// Mitsubishi GX Works2 project: 40国轩高温2次注液尝试优化   PLC: Q06UDEH (continued)

Lifter40204(ShuttleCarInOut:=LifterIO40204);	(*2线升降台*)
LifterIO40204.xCylinder:=1;
Y240:=LifterIO40204.xCW;					
Y241:=LifterIO40204.xCCW;					
LifterIO40204.xForward:=M549;					
LifterIO40204.xBackward:=M550;					
ShuttleCarCurrentPosition(X45 OR X44,X44,X45,FALSE,LifterIO40204.iCurrentPos);					
M647:=LifterIO40204.xOvertimeAlarm ;					
LifterIO40204.diDeviceID:=40204;					

Lifter40205(ShuttleCarInOut:=LifterIO40205);		(*3线升降台*)
LifterIO40205.xCylinder:=1;			
Y242:=LifterIO40205.xCW;					
Y243:=LifterIO40205.xCCW;					
LifterIO40205.xForward:=M551;					
LifterIO40205.xBackward:=M552;					
ShuttleCarCurrentPosition(X47 OR X46,X47,X46,FALSE,LifterIO40205.iCurrentPos);					
M648:=LifterIO40205.xOvertimeAlarm ;					
LifterIO40205.diDeviceID:=40205;					

Lifter40206(ShuttleCarInOut:=LifterIO40206);	(*4线升降台*)	
LifterIO40206.xCylinder:=1;			
Y276:=LifterIO40206.xCW;					
Y244:=LifterIO40206.xCCW;					
LifterIO40206.xForward:=M553;					
LifterIO40206.xBackward:=M554;					
ShuttleCarCurrentPosition(X49 OR X48,X48,X49,FALSE,LifterIO40206.iCurrentPos);					
M649:=LifterIO40206.xOvertimeAlarm ;					
LifterIO40206.diDeviceID:=40206;					

Lifter40207(ShuttleCarInOut:=LifterIO40207);	(*高温入库顶起机构*)	
LifterIO40207.xCylinder:=1;			
Y256:=LifterIO40207.xCW;					
Y257:=LifterIO40207.xCCW;					
LifterIO40207.xForward:=M556;					
LifterIO40207.xBackward:=M583;					
ShuttleCarCurrentPosition(X66 OR X65,X66,X65,FALSE,LifterIO40207.iCurrentPos);					
LifterIO40206.diDeviceID:=40207;
M651:=LifterIO40207.xOvertimeAlarm ;	

Lifter40208(ShuttleCarInOut:=LifterIO40208);	(*高温出库顶起机构*)	
LifterIO40208.xCylinder:=1;			
Y25A:=LifterIO40208.xCW;					
Y25B:=LifterIO40208.xCCW;					
LifterIO40208.xForward:=M558;					
LifterIO40208.xBackward:=M584;					
ShuttleCarCurrentPosition(X6A OR X69,X6A,X69,FALSE,LifterIO40208.iCurrentPos);					
LifterIO40206.diDeviceID:=40208;	
M653:=LifterIO40206.xOvertimeAlarm ;		

Switch40301(ConveyorEntryIO:=ConveyorIO40101 ,ConveyorExitIO:=ConveyorIO40102 ,SwitchIO:=SwitchIO40301);(*高温入库*)
SwitchIO40301.xLiftCylinderRetractDetect:=X64;							
SwitchIO40301.xLiftCylinderExtendDetect:=X63;							
Y254:=SwitchIO40301.xLiftCylinderExtend;							
SwitchIO40301.xLiftCylinderExtendButton:=M555;	
SwitchIO40301.xLiftCylinderRetractButton:=NOT M555;						
M650:=SwitchIO40301.xOvertimeAlarm ;							

(*Switch40302(ConveyorEntryIO:=ConveyorIO40103 ,ConveyorExitIO:=ConveyorIO40104 ,SwitchIO:=SwitchIO40302);*)(*高温入库里面*)(*
SwitchIO40302.xLiftCylinderRetractDetect:=X66;						
SwitchIO40302.xLiftCylinderExtendDetect:=X65;		*)										
						

Switch40303(ConveyorEntryIO:=ConveyorIO40106 ,ConveyorExitIO:=ConveyorIO40109 ,SwitchIO:=SwitchIO40303);(*高温出库*)
SwitchIO40303.xLiftCylinderExtendInit:=1;
SwitchIO40303.xLiftCylinderRetractDetect:=X68;							
SwitchIO40303.xLiftCylinderExtendDetect:=X67;							
Y258:=SwitchIO40303.xLiftCylinderExtend;							
SwitchIO40303.xLiftCylinderExtendButton:=M557;	
SwitchIO40303.xLiftCylinderRetractButton:=NOT M557;						
M652:=SwitchIO40303.xOvertimeAlarm ;							
SwitchIO40303.xLiftCylinderExtendInit:=1;

Switch40304(ConveyorEntryIO:=ConveyorIO40108 ,ConveyorExitIO:=ConveyorIO40107 ,SwitchIO:=SwitchIO40304);(*高温出库里面*)
SwitchIO40304.xLiftCylinderExtendInit:=1;
SwitchIO40304.xLiftCylinderRetractDetect:=X6A;	(*顶起部分单独写了*)						
SwitchIO40304.xLiftCylinderExtendDetect:=X69;											
SwitchIO40304.xLiftCylinderExtendInit:=1;						

Switch40305(ConveyorEntryIO:=ConveyorIO40114 ,ConveyorExitIO:=ConveyorIO40110 ,SwitchIO:=SwitchIO40305);(*1线上层*)
SwitchIO40305.xLiftCylinderRetractDetect:=X6C;							
SwitchIO40305.xLiftCylinderExtendDetect:=X6B;							
Y25C:=SwitchIO40305.xLiftCylinderExtend;							
Y270:=SwitchIO40305.xExitBarCylinderRetract;							
SwitchIO40305.xLiftCylinderExtendButton:=M559;	
SwitchIO40305.xLiftCylinderRetractButton:=NOT M559;						
SwitchIO40305.xExitBarCylinderRetractButton:=M560;							
M654:=SwitchIO40305.xOvertimeAlarm ;							

Switch40306(ConveyorEntryIO:=ConveyorIO40112 ,ConveyorExitIO:=ConveyorIO40113 ,SwitchIO:=SwitchIO40306);(*2线上层*)
SwitchIO40306.xLiftCylinderRetractDetect:=X6E;							
SwitchIO40306.xLiftCylinderExtendDetect:=X6D;							
Y25E:=SwitchIO40306.xLiftCylinderExtend;							
Y279:=SwitchIO40306.xExitBarCylinderRetract;							
SwitchIO40306.xLiftCylinderExtendButton:=M561;	
SwitchIO40306.xLiftCylinderRetractButton:=NOT M561;						
SwitchIO40306.xExitBarCylinderRetractButton:=M562;							
M655:=SwitchIO40306.xOvertimeAlarm ;							

Switch40307(ConveyorEntryIO:=ConveyorIO40115 ,ConveyorExitIO:=ConveyorIO40116 ,SwitchIO:=SwitchIO40307);(*3线上层*)
SwitchIO40307.xLiftCylinderRetractDetect:=X70;							
SwitchIO40307.xLiftCylinderExtendDetect:=X6F;							
Y260:=SwitchIO40307.xLiftCylinderExtend;							
Y27A:=SwitchIO40307.xExitBarCylinderRetract;							
SwitchIO40307.xLiftCylinderExtendButton:=M563;	
SwitchIO40307.xLiftCylinderRetractButton:=NOT M563;						
SwitchIO40307.xExitBarCylinderRetractButton:=M564;							
M656:=SwitchIO40307.xOvertimeAlarm ;							

Switch40308(ConveyorEntryIO:=ConveyorIO40118 ,ConveyorExitIO:=ConveyorIO40119 ,SwitchIO:=SwitchIO40308);(*4线上层*)
SwitchIO40308.xLiftCylinderRetractDetect:=X72;							
SwitchIO40308.xLiftCylinderExtendDetect:=X71;							
Y262:=SwitchIO40308.xLiftCylinderExtend;							
Y27B:=SwitchIO40308.xExitBarCylinderRetract;							
SwitchIO40308.xLiftCylinderExtendButton:=M565;	
SwitchIO40308.xLiftCylinderRetractButton:=NOT M565;						
SwitchIO40308.xExitBarCylinderRetractButton:=M566;							
M657:=SwitchIO40308.xOvertimeAlarm ;							

Switch40309(ConveyorEntryIO:=ConveyorIO40122 ,ConveyorExitIO:=ConveyorIO40120 ,SwitchIO:=SwitchIO40309);(*4线下层*)
SwitchIO40309.xLiftCylinderExtendInit:=1;
SwitchIO40309.xLiftCylinderRetractDetect:=X74;							
SwitchIO40309.xLiftCylinderExtendDetect:=X73;							
Y264:=SwitchIO40309.xLiftCylinderExtend;							
SwitchIO40309.xLiftCylinderExtendButton:=M567;	
SwitchIO40309.xLiftCylinderRetractButton:=NOT M567;						
M658:=SwitchIO40309.xOvertimeAlarm ;							

Switch40310(ConveyorEntryIO:=ConveyorIO40124 ,ConveyorExitIO:=ConveyorIO40126 ,SwitchIO:=SwitchIO40310);(*3线下层*)
SwitchIO40310.xLiftCylinderExtendInit:=1;
SwitchIO40310.xLiftCylinderRetractDetect:=X76;							
SwitchIO40310.xLiftCylinderExtendDetect:=X75;							
Y266:=SwitchIO40310.xLiftCylinderExtend;							
SwitchIO40310.xLiftCylinderExtendButton:=M568;		
SwitchIO40310.xLiftCylinderRetractButton:=NOT M568;					
M659:=SwitchIO40310.xOvertimeAlarm ;							

Switch40311(ConveyorEntryIO:=ConveyorIO40128 ,ConveyorExitIO:=ConveyorIO40129,SwitchIO:=SwitchIO40311);(*2线下层*)
SwitchIO40311.xLiftCylinderExtendInit:=1;
SwitchIO40311.xLiftCylinderRetractDetect:=X77;							
SwitchIO40311.xLiftCylinderExtendDetect:=X78;							
Y268:=SwitchIO40311.xLiftCylinderExtend;							
SwitchIO40311.xLiftCylinderExtendButton:=M569;	
SwitchIO40311.xLiftCylinderRetractButton:=NOT M569;						
M660:=SwitchIO40311.xOvertimeAlarm ;							

Switch40312(ConveyorEntryIO:=ConveyorIO40131 ,ConveyorExitIO:=ConveyorIO40132 ,SwitchIO:=SwitchIO40312);(*1线下层*)
SwitchIO40312.xLiftCylinderExtendInit:=1;(*先写为0，等顶升修好了再改回1*)
SwitchIO40312.xLiftCylinderRetractDetect:=X7A;							
SwitchIO40312.xLiftCylinderExtendDetect:=X79;							
Y26A:=SwitchIO40312.xLiftCylinderExtend;							
SwitchIO40312.xLiftCylinderExtendButton:=M570;
SwitchIO40312.xLiftCylinderRetractButton:=NOT M570;							
M661:=SwitchIO40312.xOvertimeAlarm ;	

(*叠盘*)
Folder40501(FolderIO:= FolderIO40501 ,FolderConveyorIO:= ConveyorIO40209);
(*夹紧气缸*)
FolderIO40501.i_xCylinderGrabExtendDetect:=X55 ;
FolderIO40501.i_xCylinderGrabRetractDetect:=X56 ;
Y250:=FolderIO40501.o_xCylinderGrabExtend;
Y251:=FolderIO40501.o_xCylinderGrabRetract;
FolderIO40501.i_xCylinderGrabExtendButton:=M571;
FolderIO40501.i_xCylinderGrabRetractButton:=M572;
(*上层气缸*)
FolderIO40501.i_xCylinderUpExtendDetect:=X54;
FolderIO40501.i_xCylinderUpRetractDetect:=X53;
Y24A:=FolderIO40501.o_xCylinderUpExtend;
Y24B:=FolderIO40501.o_xCylinderUpRetract;
FolderIO40501.i_xCylinderUpExtendButton:=M573;
FolderIO40501.i_xCylinderUpRetractButton:=M574;
(*下层气缸*)
FolderIO40501.i_xCylinderDownExtendDetect:=X52;
FolderIO40501.i_xCylinderDownRetractDetect:=X51;
Y249:=FolderIO40501.o_xCylinderDownExtend;
Y248:=FolderIO40501.o_xCylinderDownRetract;
FolderIO40501.i_xCylinderDownExtendButton:=M575;
FolderIO40501.i_xCylinderDownRetractButton:=M576;
M662:=FolderIO40501.o_xUpCylinderError;
M663:=FolderIO40501.o_xDownCylinderError;
M664:=FolderIO40501.o_xGrabCylinderError;

(*拆盘*)
DivideFolder40502(FolderIO:= DivideFolderIO40502 ,FolderConveyorIO:=ConveyorIO40105);
(*夹紧气缸*)
DivideFolderIO40502.i_xCylinderGrabExtendDetect:=X5D;
DivideFolderIO40502.i_xCylinderGrabRetractDetect:=X5E;
Y252:=DivideFolderIO40502.o_xCylinderGrabExtend;
Y253:=DivideFolderIO40502.o_xCylinderGrabRetract;
DivideFolderIO40502.i_xCylinderGrabExtendButton:=M577;
DivideFolderIO40502.i_xCylinderGrabRetractButton:=M578;
(*上层气缸*)
DivideFolderIO40502.i_xCylinderUpExtendDetect:=X5C;
DivideFolderIO40502.i_xCylinderUpRetractDetect:=X5B;
Y24E:=DivideFolderIO40502.o_xCylinderUpExtend;
Y24F:=DivideFolderIO40502.o_xCylinderUpRetract;
DivideFolderIO40502.i_xCylinderUpExtendButton:=M579;
DivideFolderIO40502.i_xCylinderUpRetractButton:=M580;
(*下层气缸*)
DivideFolderIO40502.i_xCylinderDownExtendDetect:=X5A;
DivideFolderIO40502.i_xCylinderDownRetractDetect:=X59;
Y24C:=DivideFolderIO40502.o_xCylinderDownExtend;
Y24D:=DivideFolderIO40502.o_xCylinderDownRetract;
DivideFolderIO40502.i_xCylinderDownExtendButton:=M581;
DivideFolderIO40502.i_xCylinderDownRetractButton:=M582;
M665:=DivideFolderIO40502.o_xUpCylinderError;
M666:=DivideFolderIO40502.o_xDownCylinderError;
M667:=DivideFolderIO40502.o_xGrabCylinderError;
			
(*******************上位机通信数据*******************************)
(*扫码位，虚拟的*)
ComConveyor40140(ConveyorIO:=ConveyorIO40140,CommunicationIO:=ComConveyorIO40140);
ComConveyorIO40140.i_iResponsPCPLC:=D2000;	
ComConveyorIO40140.i_iTypeInfoPCPLC:=D2001;
ComConveyorIO40140.i_iReadWriteFlagPCPLC:=D2005;	
ComConveyorIO40140.i_iTaskProcessFlagPCPLC:=D2006;	
ComConveyorIO40140.i_iCommandPCPLC:=D2007;	
ComConveyorIO40140.i_iTaskIDPCPLC:=D2008;	
DMOV(TRUE,D2009,ComConveyorIO40140.i_diDestinationDevicePCPLC);	
ComConveyorIO40140.i_iProductIDPCPLC:=D2011;	
D3000:=ComConveyorIO40140.o_iRequestPLCPC;	
D3001:=ComConveyorIO40140.o_iForceInportPLCPC;
D3002:=ComConveyorIO40140.o_iFolderNumberPLCPC;
D3003:=ComConveyorIO40140.o_iEmptyPLCPC;
D3005:=ComConveyorIO40140.o_iReadWriteFlagPLCPC;	
D3006:=ComConveyorIO40140.o_iDeviceStatusPLCPC;	
D3007:=ComConveyorIO40140.o_iTaskIDPLCPC;	
D3008:=ComConveyorIO40140.o_iProductIDPLCPC;	
ComConveyorIO40140.i_xExportConveyor:=0;
(*碟盘位*)
ComConveyor40209(ConveyorIO:=ConveyorIO40209,CommunicationIO:=ComConveyorIO40209);
ComConveyorIO40209.i_iResponsPCPLC:=D2015;	
ComConveyorIO40209.i_iTypeInfoPCPLC:=D2016;
ComConveyorIO40209.i_iReadWriteFlagPCPLC:=D2020;	
ComConveyorIO40209.i_iTaskProcessFlagPCPLC:=D2021;	
ComConveyorIO40209.i_iCommandPCPLC:=D2022;	
ComConveyorIO40209.i_iTaskIDPCPLC:=D2023;	
DMOV(TRUE,D2024,ComConveyorIO40209.i_diDestinationDevicePCPLC);	
ComConveyorIO40209.i_iProductIDPCPLC:=D2026;	
D3015:=ComConveyorIO40209.o_iRequestPLCPC;	
D3016:=ComConveyorIO40209.o_iForceInportPLCPC;
D3017:=ComConveyorIO40209.o_iFolderNumberPLCPC;
D3018:=ComConveyorIO40209.o_iEmptyPLCPC;
D3020:=ComConveyorIO40209.o_iReadWriteFlagPLCPC;	
D3021:=ComConveyorIO40209.o_iDeviceStatusPLCPC;	
D3022:=ComConveyorIO40209.o_iTaskIDPLCPC;	
D3023:=ComConveyorIO40209.o_iProductIDPLCPC;	
(*入库1站台*)
ComConveyor40111(ConveyorIO:=ConveyorIO40111,CommunicationIO:=ComConveyorIO40111);
ComConveyorIO40111.i_iResponsPCPLC:=D2030;	
ComConveyorIO40111.i_iTypeInfoPCPLC:=D2031;
ComConveyorIO40111.i_iReadWriteFlagPCPLC:=D2035;	
ComConveyorIO40111.i_iTaskProcessFlagPCPLC:=D2036;	
ComConveyorIO40111.i_iCommandPCPLC:=D2037;	
ComConveyorIO40111.i_iTaskIDPCPLC:=D2038;	
DMOV(TRUE,D2039,ComConveyorIO40111.i_diDestinationDevicePCPLC);	
ComConveyorIO40111.i_iProductIDPCPLC:=D2041;	
D3030:=ComConveyorIO40111.o_iRequestPLCPC;	
D3031:=ComConveyorIO40111.o_iForceInportPLCPC;
D3032:=ComConveyorIO40111.o_iFolderNumberPLCPC;
D3033:=ComConveyorIO40111.o_iEmptyPLCPC;
D3035:=ComConveyorIO40111.o_iReadWriteFlagPLCPC;	
D3036:=ComConveyorIO40111.o_iDeviceStatusPLCPC;	
D3037:=ComConveyorIO40111.o_iTaskIDPLCPC;	
D3038:=ComConveyorIO40111.o_iProductIDPLCPC;	
(*入库2站台*)
ComConveyor40104(ConveyorIO:=ConveyorIO40104,CommunicationIO:=ComConveyorIO40104);
ComConveyorIO40104.i_iResponsPCPLC:=D2045;	
ComConveyorIO40104.i_iTypeInfoPCPLC:=D2046;
ComConveyorIO40104.i_iReadWriteFlagPCPLC:=D2050;	
ComConveyorIO40104.i_iTaskProcessFlagPCPLC:=D2051;	
ComConveyorIO40104.i_iCommandPCPLC:=D2052;	
ComConveyorIO40104.i_iTaskIDPCPLC:=D2053;	
DMOV(TRUE,D2054,ComConveyorIO40104.i_diDestinationDevicePCPLC);	
ComConveyorIO40104.i_iProductIDPCPLC:=D2056;	
D3045:=ComConveyorIO40104.o_iRequestPLCPC;
D3046:=ComConveyorIO40104.o_iForceInportPLCPC;
D3047:=ComConveyorIO40104.o_iFolderNumberPLCPC;
IF D3045=2 THEN
	D3048:=ComConveyorIO40104.o_iEmptyPLCPC;
ELSE
	D3048:=1;
END_IF;	
D3050:=ComConveyorIO40104.o_iReadWriteFlagPLCPC;	
D3051:=ComConveyorIO40104.o_iDeviceStatusPLCPC;	
D3052:=ComConveyorIO40104.o_iTaskIDPLCPC;	
D3053:=ComConveyorIO40104.o_iProductIDPLCPC;	(*XB是紧挨着入库口1那个开关，顶起之后，再运一会儿，运到这个开关才发请求*)
ComConveyorIO40104.i_xExtraCondition:=LifterIO40207.iCurrentPos=2 AND NOT m_xImport  AND XB; 
(*出库1站台*)
ComConveyor40105(ConveyorIO:=ConveyorIO40105,CommunicationIO:=ComConveyorIO40105);
ComConveyorIO40105.i_iResponsPCPLC:=D2060;	
ComConveyorIO40105.i_iTypeInfoPCPLC:=D2061;
ComConveyorIO40105.i_iReadWriteFlagPCPLC:=D2065;	
ComConveyorIO40105.i_iTaskProcessFlagPCPLC:=D2066;	
ComConveyorIO40105.i_iCommandPCPLC:=D2067;	
ComConveyorIO40105.i_iTaskIDPCPLC:=D2068;	
DMOV(TRUE,D2069,ComConveyorIO40105.i_diDestinationDevicePCPLC);	
ComConveyorIO40105.i_iProductIDPCPLC:=D2071;	
D3060:=ComConveyorIO40105.o_iRequestPLCPC;	
D3061:=ComConveyorIO40105.o_iForceInportPLCPC;
D3062:=ComConveyorIO40105.o_iFolderNumberPLCPC;
D3063:=ComConveyorIO40105.o_iEmptyPLCPC;
D3065:=ComConveyorIO40105.o_iReadWriteFlagPLCPC;	
D3066:=ComConveyorIO40105.o_iDeviceStatusPLCPC;	
D3067:=ComConveyorIO40105.o_iTaskIDPLCPC;	
D3068:=ComConveyorIO40105.o_iProductIDPLCPC;	
ComConveyorIO40105.i_xExportConveyor:=1;
ComConveyorIO40105.i_xExtraCondition:=ConveyorIO40107.xEmpty AND NOT ConveyorIO40108.xCWPresent  AND NOT ConveyorIO40107.xCWPresent 
																						AND LifterIO40208.iCurrentPos=2 AND X69
																						AND NOT g_x36HourExport1Forbidden;(*无出库禁止*)

(*******************以上是上位机通信数据*******************************)

	(*数据传递*)
	ConveyorIO40209.diDesConveyorIn:=ConveyorIO40140.diDesConveyorOut;
	ConveyorIO40209.iTaskIDIn:=ConveyorIO40140.iTaskIDOut;
	ConveyorIO40209.iProductCategoryIn:=ConveyorIO40209.iProductCategoryOut;
	ConveyorIO40101.diDesConveyorIn:=ConveyorIO40140.diDesConveyorOut(*ConveyorIO40209.diDesConveyorOut*);
	ConveyorIO40101.iTaskIDIn:=ConveyorIO40140.iTaskIDOut(*ConveyorIO40209.iTaskIDOut*);
	ConveyorIO40101.iProductCategoryIn:=ConveyorIO40140.iProductCategoryOut;
	IF ConveyorIO40102.diDesConveyorOut>0 THEN		
		ConveyorIO401021.diDesConveyorIn:=ConveyorIO40102.diDesConveyorOut;
		ConveyorIO401021.iTaskIDIn:=ConveyorIO40102.iTaskIDOut;
		ConveyorIO401021.iProductCategoryIn:=ConveyorIO40102.iProductCategoryOut;
	END_IF;
	ConveyorIO40103.diDesConveyorIn:=ConveyorIO401021.diDesConveyorOut;
	ConveyorIO40103.iTaskIDIn:=ConveyorIO401021.iTaskIDOut;
	ConveyorIO40103.iProductCategoryIn:=ConveyorIO401021.iProductCategoryOut;
	ConveyorIO40104.diDesConveyor:=ConveyorIO40103.diDesConveyor;
	ConveyorIO40104.iTaskID:=ConveyorIO40103.iTaskID;
	ConveyorIO40104.iProductCategory:=ConveyorIO40103.iProductCategory;
	ConveyorIO40111.diDesConveyorIn:=ConveyorIO40104.diDesConveyorOut;
	ConveyorIO40111.iTaskIDIn:=ConveyorIO40104.iTaskIDOut;
	ConveyorIO40111.iProductCategoryIn:=ConveyorIO40104.iProductCategoryOut;		
	(*自动部分*)
IF g_xAuto THEN
(*	D221.4:=FolderIO40501.o_xEntryPermit AND ConveyorIO40101.xEmpty;
	FolderIO40501.i_xEntryEnable:=D421.4;
	FolderIO40501.i_xExitEnable:=ConveyorIO40101.xEmpty;*)(*临时不叠盘，直接过*)
	D221.4:=ConveyorIO40101.xEmpty AND ConveyorIO40140.xNextRun(*这个是30线体的Unload信号*);
							(*AND FolderIO40501.o_xEntryPermit;*)
	ConveyorIO40140.xLoad:=D421.5;
	D221.5:=ConveyorIO40140.xNextRun;
	dmov(ConveyorIO40140.xEmpty,0,ConveyorIO40140.diDesConveyor);(*_以前走load流程，不需要这个，现在走putinto，就需要了_*)
	ConveyorIO40140.xUnload:=ConveyorIO40101.xEmpty AND ConveyorIO40140.diDesConveyor<>0;
															(*AND FolderIO40501.o_xEntryPermit ;
		FolderIO40501.i_xEntryEnable:=D421.4 OR M8;*)(*这个是30那边的NextRun*)
	(*FolderIO40501.i_xExitEnable:=ConveyorIO40101.xEmpty;*)
	
	
	SwitchIO40301.xEntryEnable:=D421.4 OR M8 OR ConveyorIO40140.xNextRun(*屏蔽碟盘*);
	SwitchIO40301.xSwithEnable:=1;
	SwitchIO40301.xExitEnable:= ConveyorIO401021.xEmpty;
	ConveyorIO401021.xLoad:=ConveyorIO40102.xNextRun;
	ConveyorIO401021.xUnload:=ConveyorIO40103.xEmpty 
																(*AND LifterIO40201.iCurrentPos=2 AND X3F*)
																AND LifterIO40207.iCurrentPos=1 AND X66
																AND(ConveyorIO401021.diDesConveyor=40104(*目标是40104时不需要额外条件*)
																			OR(ConveyorIO401021.diDesConveyor=40111 AND  ConveyorIO40111.xEmpty AND ConveyorIO40104.xEmpty)); 
																			(*目标是40111时，如果有一个正在往40111送，也不下料*)
(*强制入库，如果连续两个都是去40111，那么强制入库*)
IF NOT ConveyorIO401021.xEmpty AND ConveyorIO401021.diDesConveyor=40111 AND NOT ConveyorIO40111.xEmpty AND ConveyorIO40103.xEmpty  
			OR g_xForceImport		THEN 
		 ComConveyorIO40111.o_iForceInportPLCPC:=2;
	ELSE
		 ComConveyorIO40111.o_iForceInportPLCPC:=1;
END_IF;
	IF ConveyorIO40104.xEmpty AND ConveyorIO40111.xEmpty THEN
		g_xForceImport:=0;
	END_IF;	
	
	(*高温入库门控制*)
	IF NOT ConveyorIO401021.xEmpty AND ConveyorIO40103.xEmpty THEN
		LifterIO40201.xMDIExe:=1;
		LifterIO40201.iDestinationPos:=2;
	ELSE
		LifterIO40201.xMDIExe:=1;
		LifterIO40201.iDestinationPos:=1;
	END_IF;	
	ConveyorIO40103.xLoad:=ConveyorIO401021.xNextRun;
	(*X66是末端顶起机构没顶起时的磁开关*)
	IF X66 AND LDP(TRUE,NOT ConveyorIO40103.xEmpty) AND ConveyorIO40104.xCWPresent THEN(*入线体刷新顶升线体,在进来时才刷*)
		ConveyorIO40104.xPutInto:=1;
	ELSIF LDP(TRUE,NOT ConveyorIO40104.xEmpty) THEN
		ConveyorIO40104.xPutInto:=0;
	END_IF;	
	IF LDP(TRUE,ConveyorIO40104.xEmpty)THEN(*顶升线体刷新入线体*)
		ConveyorIO40103.xPutInto:=1;
	ELSIF 	 LDP(TRUE,ConveyorIO40103.xEmpty)THEN
		ConveyorIO40103.xPutInto:=0;
	END_IF;
	(*顶升部分单独写，防止用switch意外顶翻料框*)
	LifterIO40207.xMDIExe:=1;(*本来打算直接开关控制MDIexe，但MDI信号一没，就会往下降，会有问题，所以开关改到目标地址里面了*)
	(*NOT ConveyorIO40103.xError AND NOT ConveyorIO40111.xError;*)(*这里打算不用线体error了，因为线体error会不好复位*)
	IF NOT ConveyorIO40104.xEmpty AND NOT X6 THEN(*升起必须连框开关没挡住*)
		LifterIO40207.iDestinationPos:=2;
	ELSIF ConveyorIO40104.xEmpty AND NOT XB THEN(*下降需中间开关没挡住*)
		LifterIO40207.iDestinationPos:=1;
	END_IF;
	ConveyorIO40104.xUnload:=ConveyorIO40111.xEmpty 
															AND LifterIO40207.iCurrentPos=2 AND X65
															AND ConveyorIO40104.diDesConveyor=40111;	
	ConveyorIO40111.xLoad:=ConveyorIO40104.xNextRun;(*这是40104下料给40111的，还需要写一个40104上到位自己转的*)
	(*这里顶起来了之后，多转3S，让他到位*)
	m_TonImportDelay(IN:= m_xImport,PT:=t#3S,Q:= m_xImportDelay ,ET:= m_tImportDelay );
	IF LDP(TRUE,LifterIO40207.iCurrentPos=2)AND NOT ConveyorIO40104.xEmpty THEN
		m_xImport:=1;
	ELSIF  m_xImportDelay THEN
		m_xImport:=0;
	END_IF;	

	
	ConveyorIO40111.xPutInto:=SM413 AND NOT ConveyorIO40111.xBusy;
	IF LifterIO40207.iCurrentPos=2 AND X65 THEN
		SET(LDP(TRUE, ConveyorIO40111.xPutInto) , ConveyorIO40104.xPutInto);
		RST(LDF(TRUE, ConveyorIO40111.xPutInto) , ConveyorIO40104.xPutInto);		
		RST(ConveyorIO40104.xEmpty , ConveyorIO40104.xPutInto);
	END_IF;
	(*线体的putinto信号在通信块里写好了，所以这里就不写了。*)
	OUT_T( ConveyorIO40108.xCWPresent AND NOT ConveyorIO40108.xBusy
					 AND LifterIO40208.iCurrentPos=2 AND ConveyorIO40108.xEmpty,
						 TC5 , 100 );
	ConveyorIO40105.xPutInto:=TS5 ;(*触摸屏做一个送完刷新按钮，到时候上位机控制*)
	IF LDP(TRUE,ConveyorIO40105.xPutInto)THEN
		ConveyorIO40108.xPutInto:=1;(*这里直接:=不行，因为108还是switch的一部分，会导致switch里的putinto无法生效*)
	ELSIF LDF(TRUE,ConveyorIO40105.xPutInto)	THEN
		ConveyorIO40108.xPutInto:=0;
	END_IF;	
		m_TonExportDelay(IN:= m_xExport,PT:=t#6S,Q:= m_xExportDelay ,ET:= m_tExportDelay );
	IF LifterIO40208.iCurrentPos=2 AND LDP(TRUE, NOT ConveyorIO40108.xEmpty AND NOT ConveyorIO40108.xLoad ) 
		OR ldp(TRUE,M30) THEN(*M30是触摸屏上的手动出库按钮，手动出的库需要按这个按钮*)
		m_xExport:=1;
	ELSIF  m_xExportDelay THEN
		m_xExport:=0;
	END_IF;	
	
	
	ConveyorIO40105.xUnload:=ConveyorIO40108.xEmpty AND LifterIO40208.iCurrentPos=2 AND X69;
	(*顶升部分单独写，防止用switch意外顶翻料框*)
	LifterIO40208.xMDIExe:=1;
	IF ConveyorIO40108.xEmpty THEN
		LifterIO40208.iDestinationPos:=2;
	ELSIF NOT ConveyorIO40108.xEmpty AND NOT m_xExport AND NOT X7C  AND ConveyorIO401061.xEmpty THEN
		LifterIO40208.iDestinationPos:=1;		
	END_IF;	
	SwitchIO40304.xEntryEnable:=ConveyorIO40105.xNextRun;
	SwitchIO40304.xSwithEnable:=1;
	SwitchIO40304.xExitEnable:=ConveyorIO401061.xEmpty;
	ConveyorIO401061.xLoad:=ConveyorIO40107.xNextRun;
	 ConveyorIO401061.xUnload:=ConveyorIO40106.xEmpty (*AND LifterIO40202.iCurrentPos=2*);
	 
	 (*高温出库门控制*)
	IF ConveyorIO40106.xEmpty AND NOT ConveyorIO401061.xEmpty THEN
		LifterIO40202.xMDIExe:=1;
		LifterIO40202.iDestinationPos:=2;
	ELSE
		LifterIO40202.xMDIExe:=1;
		LifterIO40202.iDestinationPos:=1;
	END_IF;	
	SwitchIO40303.xEntryEnable:=ConveyorIO401061.xNextRun;
	SwitchIO40303.xSwithEnable:=1;
	SwitchIO40303.xExitEnable:=ConveyorIO40114.xEmpty ;
	(*DivideFolderIO40502.o_xEntryPermit;
	DivideFolderIO40502.i_xEntryEnable:=ConveyorIO40109.xNextRun;
	DivideFolderIO40502.i_xExitEnable:=*)(*暂时不用拆盘*)
	(*******4个位置的要料请求，排队处理********)(*——这里改掉，不在这里排队，去入库口抢占
	Task40105(	arrxCondition:=TaskCondition40105,
						xTaskComplete:=LDP(TRUE,ConveyorIO40109.xEmpty),
						xReSET:=g_xResetSingle AND g_diDeviceIDSelect=40109,
						iPriority:=m_iTask40105);
	TaskCondition40105[1].xCondition:=	ConveyorIO401191.xEmpty AND m_xLoadPermit[4];
	TaskCondition40105[2].xCondition:=	ConveyorIO401161.xEmpty AND m_xLoadPermit[3];
	TaskCondition40105[3].xCondition:=	ConveyorIO401131.xEmpty AND m_xLoadPermit[2];
	TaskCondition40105[4].xCondition:=	ConveyorIO401101.xEmpty AND m_xLoadPermit[1];
*)
(*//根据任务生成目标地址	*)(*
	DMOV(m_iTask40105=1,	40119,	ConveyorIO40109.diDesConveyor);
	DMOV(m_iTask40105=2,	40116,	ConveyorIO40109.diDesConveyor);
	DMOV(m_iTask40105=3,	40113,	ConveyorIO40109.diDesConveyor);
	DMOV(m_iTask40105=4,	40110,	ConveyorIO40109.diDesConveyor);	*)
	(*任务目标地址的传递*)
	ConveyorIO40109.diDesConveyor:=40110;(*这样控制1线阻挡进料时顶起*)
	ConveyorIO40114.diDesConveyorIn:=	ConveyorIO40109.diDesConveyorOut;
	ConveyorIO40112.diDesConveyorIn:=	ConveyorIO40114.diDesConveyorOut;
	ConveyorIO40115.diDesConveyorIn:=	ConveyorIO40112.diDesConveyorOut;
	ConveyorIO40118.diDesConveyorIn:=	ConveyorIO40115.diDesConveyorOut;
	m_xLoadPermit[1]:=M52;
	m_xLoadPermit[2]:=M53;
	m_xLoadPermit[3]:=M54;
	m_xLoadPermit[4]:=M55;
(*1线顶升排队*)	
	TaskSwitch40305(xCondition:=TaskCondition40305,
										xTaskComplete:=LDP(TRUE,ConveyorIO40114.xEmpty),
										xReset:=g_xResetSingle AND g_diDeviceIDSelect=40114,
										iPriority:= m_iTask40305 );
	TaskCondition40305[1]:=ConveyorIO40112.xEmpty;
	TaskCondition40305[2]:=ConveyorIO401101.xEmpty AND m_xLoadPermit[1];
	DMOV(m_iTask40305=1,	40113,	ConveyorIO40114.diDesConveyor);(*这么改可以控制2线出阻挡*)	
	DMOV(m_iTask40305=2,	40110,	ConveyorIO40114.diDesConveyor);(*这么改可以控制1线出阻挡顶起*)
(*2线顶升排队*)		
	TaskSwitch40306(xCondition:=TaskCondition40306,
										xTaskComplete:=LDP(TRUE,ConveyorIO40112.xEmpty),
										xReset:=g_xResetSingle AND g_diDeviceIDSelect=40112,
										iPriority:= m_iTask40306 );
	TaskCondition40306[1]:=ConveyorIO40115.xEmpty;
	TaskCondition40306[2]:=ConveyorIO401131.xEmpty AND m_xLoadPermit[2];
	DMOV(m_iTask40306=1,	40116,	ConveyorIO40112.diDesConveyor);
	DMOV(m_iTask40306=2,	40113,	ConveyorIO40112.diDesConveyor);	
(*3线顶升排队*)			
	TaskSwitch40307(xCondition:=TaskCondition40307,
										xTaskComplete:=LDP(TRUE,ConveyorIO40115.xEmpty),
										xReset:=g_xResetSingle AND g_diDeviceIDSelect=40115,
										iPriority:= m_iTask40307 );
	TaskCondition40307[1]:=ConveyorIO40118.xEmpty;
	TaskCondition40307[2]:=ConveyorIO401161.xEmpty AND m_xLoadPermit[3];
	(*DMOV(m_iTask40307=1,	40119,	ConveyorIO40115.diDesConveyor);先屏蔽掉，免得往4线送，需要再开起来*)
	DMOV(m_iTask40307=2,	40116,	ConveyorIO40115.diDesConveyor);
		
	SwitchIO40305.xEntryEnable:=ConveyorIO40109.xNextRun;
	SwitchIO40305.xSwithEnable:=ConveyorIO40114.diDesConveyor=40110;
	SwitchIO40305.xExitEnable:=(SwitchIO40305.xSwithEnable AND ConveyorIO401101.xEmpty)
															OR (NOT SwitchIO40305.xSwithEnable AND ConveyorIO40112.xEmpty);
	ConveyorIO401101.xLoad:=ConveyorIO40110.xNextRun;
	IF LDP(TRUE,NOT ConveyorIO401101.xEmpty) THEN
		m_xPickStrat[1]:=1;
	ELSIF m_xPickDone[1] OR ConveyorIO401101.xEmpty THEN
		m_xPickStrat[1]:=0;
	END_IF;
	IF g_xPickOver[1] THEN
		m_xPickDone[1]:=1;
	ELSIF ConveyorIO401101.xEmpty THEN	
		m_xPickDone[1]:=0;
	END_IF;
	
	SwitchIO40306.xEntryEnable:=ConveyorIO40114.xNextRun;
	SwitchIO40306.xSwithEnable:=ConveyorIO40112.diDesConveyor=40113;
	SwitchIO40306.xExitEnable:=(SwitchIO40306.xSwithEnable AND ConveyorIO401131.xEmpty)
															OR (NOT SwitchIO40306.xSwithEnable AND ConveyorIO40115.xEmpty);
	ConveyorIO401131.xLoad:=ConveyorIO40113.xNextRun;
	IF LDP(TRUE,NOT ConveyorIO401131.xEmpty) THEN
		m_xPickStrat[2]:=1;
	ELSIF m_xPickDone[2] OR ConveyorIO401131.xEmpty THEN
		m_xPickStrat[2]:=0;
	END_IF;
	IF g_xPickOver[2] THEN
		m_xPickDone[2]:=1;
	ELSIF ConveyorIO401131.xEmpty THEN	
		m_xPickDone[2]:=0;
	END_IF;
			
	SwitchIO40307.xEntryEnable:=ConveyorIO40112.xNextRun;
	SwitchIO40307.xSwithEnable:=ConveyorIO40115.diDesConveyor=40116;
	SwitchIO40307.xExitEnable:=(SwitchIO40307.xSwithEnable AND ConveyorIO401161.xEmpty)
															OR (NOT SwitchIO40307.xSwithEnable AND ConveyorIO40118.xEmpty);
	ConveyorIO401161.xLoad:=ConveyorIO40116.xNextRun;	
		IF LDP(TRUE,NOT ConveyorIO401161.xEmpty) THEN
			m_xPickStrat[3]:=1;
		ELSIF m_xPickDone[3] OR ConveyorIO401161.xEmpty THEN
			m_xPickStrat[3]:=0;
		END_IF;
	IF g_xPickOver[3] THEN
		m_xPickDone[3]:=1;
	ELSIF ConveyorIO401161.xEmpty THEN	
		m_xPickDone[3]:=0;
	END_IF;	
		
	SwitchIO40308.xEntryEnable:=ConveyorIO40115.xNextRun;
	SwitchIO40308.xSwithEnable:=1;
	SwitchIO40308.xExitEnable:=ConveyorIO401191.xEmpty;	
	ConveyorIO401191.xLoad:=ConveyorIO40119.xNextRun;	
		IF LDP(TRUE,NOT ConveyorIO401191.xEmpty) THEN
			m_xPickStrat[4]:=1;
		ELSIF m_xPickDone[4] OR ConveyorIO401191.xEmpty THEN
			m_xPickStrat[4]:=0;
		END_IF;
	IF g_xPickOver[4] THEN
		m_xPickDone[4]:=1;
	ELSIF ConveyorIO401191.xEmpty THEN	
		m_xPickDone[4]:=0;
	END_IF;
			
(*至此，料已运到每个注液的地方，等待对方发信号，就可以升降机动作，来运走空框了*)

(*4送出*)
	ConveyorIO401191.xUnload:=ConveyorIO40135.xEmpty 
															AND LifterIO40206.iCurrentPos=2 AND X48 (*升降台在上面*)
															AND m_xPickDone[4];(*机械手给捡完信号*)
	LifterIO40206.xMDIExe:=NOT ConveyorIO40135.xError AND NOT ConveyorIO401191.xError AND NOT ConveyorIO40122.xError;
	IF ConveyorIO40135.xEmpty THEN
		LifterIO40206.iDestinationPos:=2;
	ELSE
		LifterIO40206.iDestinationPos:=1;
	END_IF;		
	ConveyorIO40135.xLoad:=ConveyorIO401191.xNextRun;
	ConveyorIO40135.xUnload:=ConveyorIO40122.xEmpty AND LifterIO40206.iCurrentPos=1 AND X49;
	ConveyorIO40135.xUnloadCCW:=1;
	SwitchIO40309.xEntryEnable:=ConveyorIO40135.xNextRun;
	SwitchIO40309.xSwithEnable:=1;
	SwitchIO40309.xExitEnable:=ConveyorIO40129.xEmpty(*防止和3线出料冲突，所以加上busy信号*)
											 AND NOT ConveyorIO40124.xbusy;
	ConveyorIO40126.xLoad:=ConveyorIO40120.xNextRun;
	(*顶升降下去，防止卡住*)
	IF LDP(TRUE,ConveyorIO40120.xNextRun )THEN
		SwitchIO40310.xLiftCylinderExtend:=0;
		SwitchIO40310.xLiftCylinderRetract:=1;
	END_IF;
	(*给上putinto，进入switch正常流程*)
	IF LDP(TRUE,NOT ConveyorIO40126.xEmpty)AND ConveyorIO40124.xEmpty THEN
		ConveyorIO40124.xPutInto:=1;
	ELSIF LDP(TRUE,NOT ConveyorIO40124.xEmpty) THEN
		ConveyorIO40124.xPutInto:=0;
	END_IF;		
	(*送出到3线横向那里了*)

(*3送出*)
	ConveyorIO401161.xUnload:=ConveyorIO40136.xEmpty AND LifterIO40205.iCurrentPos=2 AND X46 AND m_xPickDone[3];
	ConveyorIO40136.xLoad:=ConveyorIO401161.xNextRun;
	LifterIO40205.xMDIExe:=NOT ConveyorIO40136.xError AND NOT ConveyorIO401161.xError AND NOT ConveyorIO40124.xError;
	(*升降台控制*)
	IF ConveyorIO40136.xEmpty THEN
		LifterIO40205.iDestinationPos:=2;
	ELSE
		LifterIO40205.iDestinationPos:=1;
	END_IF;		
	(*这里就不做抢占任务了，在下料条件里加上not busy信号得了*)
	(*36是升降台*)(*24是下层线体*)(*26是2线下层线体*)
	ConveyorIO40136.xUnload:=ConveyorIO40124.xEmpty AND LifterIO40205.iCurrentPos=1 AND X47
														AND  NOT ConveyorIO40126.xBusy;(*未处于运行状态，表示没有在执行任务*)
	ConveyorIO40136.xUnloadCCW:=1;
	SwitchIO40310.xEntryEnable:=ConveyorIO40136.xNextRun;
	SwitchIO40310.xSwithEnable:=1;
	SwitchIO40310.xExitEnable:=ConveyorIO40129.xEmpty(*防止和2线出料冲突，所以加上busy信号*)
											 AND NOT ConveyorIO40128.xbusy;
	ConveyorIO40129.xLoad:=ConveyorIO40126.xNextRun;
	(*顶升下去，防止卡住*)
	IF LDP(TRUE,ConveyorIO40126.xNextRun )THEN
		SwitchIO40311.xLiftCylinderExtend:=0;
		SwitchIO40311.xLiftCylinderRetract:=1;
	END_IF;
	(*给上putinto，进入switch正常流程*)
	IF LDP(TRUE,NOT ConveyorIO40129.xEmpty) AND ConveyorIO40128.xEmpty THEN(*这不加个empty会出问题，正常流程也会置位putinto，而且不复位*)
		ConveyorIO40128.xPutInto:=1;
	ELSIF LDP(TRUE,NOT ConveyorIO40128.xEmpty) THEN
		ConveyorIO40128.xPutInto:=0;
	END_IF;		
	(*送出到2线横向那里了*)
